// TIA Portal project "EMS" (V15.1) (continued)
   "Carrier_08_G120DStatusWord.3" AT %I762.3 : Bool;   // Bit_03_FAULT
   "Carrier_08_G120DStatusWord.4" AT %I762.4 : Bool;   // Bit_04_OFF2
   "Carrier_08_G120DStatusWord.5" AT %I762.5 : Bool;   // Bit_05_OFF3
   "Carrier_08_G120DStatusWord.6" AT %I762.6 : Bool;   // Bit_06_LOCK_OUT
   "Carrier_08_G120DStatusWord.7" AT %I762.7 : Bool;   // Bit_07_WARN
   "Carrier_08_G120DStatusWord.8" AT %I763.0 : Bool;   // Bit_08_NO_DEVIATION
   "Carrier_08_G120DStatusWord.9" AT %I763.1 : Bool;   // Bit_09_CONTR_PLC
   "Carrier_08_G120DStatusWord.10" AT %I763.2 : Bool;   // Bit_10_F_MAX
   "Carrier_08_G120DStatusWord.11" AT %I763.3 : Bool;   // Bit_11_LIMIT_REACHED
   "Carrier_08_G120DStatusWord.12" AT %I763.4 : Bool;   // Bit_12_BRAKE_OPEN
   "Carrier_08_G120DStatusWord.13" AT %I763.5 : Bool;   // Bit_13_NO_OVERTEMP
   "Carrier_08_G120DStatusWord.14" AT %I763.6 : Bool;   // Bit_14_CW_CCW
   "Carrier_08_G120DStatusWord.15" AT %I763.7 : Bool;   // Bit_15_OVERL
   "Carrier_08_Slot2_Input" AT %IW764 : Word;   // SLOT 2 INPUT WORD
   "Carrier_08_CrashDetectSW" AT %I764.0 : Bool;   // CRASH DETECT SW
   "Carrier_08_SpareSafetyInput(2_1)" AT %I764.1 : Bool;   // SPARE SAFETY INPUT
   "Carrier_08_SpareSafetyInput(2_2)" AT %I764.2 : Bool;   // SPARE SAFETY INPUT
   "Carrier_08_SpareSafetyInput(2_3)" AT %I764.3 : Bool;   // SPARE SAFETY INPUT
   "Carrier_08_SpareSafetyInput(2_4)" AT %I764.4 : Bool;   // SPARE SAFETY INPUT
   "Carrier_08_SpareSafetyInput(2_5)" AT %I764.5 : Bool;   // SPARE SAFETY INPUT
   "Carrier_08_SpareSafetyInput(2_6)" AT %I764.6 : Bool;   // SPARE SAFETY INPUT
   "Carrier_08_SpareSafetyInput(2_7)" AT %I764.7 : Bool;   // SPARE SAFETY INPUT
   "Carrier_08_Slot3_SafetyOutput" AT %IW765 : Word;   // SLOT 3 SAFETY OUTPUT WORD
   "Carrier_08_Crash_Detect_OK" AT %I765.0 : Bool;   // CARRIER CRASH DETECT
   "Carrier_08_SpareSafetyOutput(3_1)" AT %I765.1 : Bool;   // SPARE SAFETY OUTPUT
   "Carrier_08_SpareSafetyOutput(3_2)" AT %I765.2 : Bool;   // SPARE SAFETY OUTPUT
   "Carrier_08_SpareSafetyOutput(3_3)" AT %I765.3 : Bool;   // SPARE SAFETY OUTPUT
   "Carrier_08_SpareSafetyOutput(3_4)" AT %I765.4 : Bool;   // SPARE SAFETY OUTPUT
   "Carrier_08_SpareSafetyOutput(3_5)" AT %I765.5 : Bool;   // SPARE SAFETY OUTPUT
   "Carrier_08_SpareSafetyOutput(3_6)" AT %I765.6 : Bool;   // SPARE SAFETY OUTPUT
   "Carrier_08_SpareSafetyOutput(3_7)" AT %I765.7 : Bool;   // SPARE SAFETY OUTPUT
   "Carrier_08_Slot4_Input" AT %IW766 : Word;   // SLOT 4 INPUT WORD
   "Carrier_08_480VPowerOn_MDCB1" AT %I766.0 : Bool;   // 480 VAC POWER ON MDCB 1
   "Carrier_08_SpareInput(4_1)" AT %I766.1 : Bool;   // SPARE INPUT
   "Carrier_08_SpareInput(4_2)" AT %I766.2 : Bool;   // SPARE INPUT
   "Carrier_08_SitopSelectStatus" AT %I766.3 : Bool;   // SITOP SELECT STATUS
   "Carrier_08_DCsupplyOnPSCB2" AT %I766.4 : Bool;   // DC SUPPLY ON PSCB 2
   "Carrier_08_SpareInput(4_5)" AT %I766.5 : Bool;   // SPARE INPUT
   "Carrier_08_SpareInput(4_6)" AT %I766.6 : Bool;   // SPARE INPUT
   "Carrier_08_SpareInput(4_7)" AT %I766.7 : Bool;   // SPARE INPUT
   "Carrier_08_PB1_ProdHoldLH" AT %I767.0 : Bool;   // PB 1 PRODUCTION HOLD LH
   "Carrier_08_PB2_ResetLH" AT %I767.1 : Bool;   // PB 2 RESET LH
   "Carrier_08_PB3_ProdHoldRH" AT %I767.2 : Bool;   // PB 3 PRODUCTION HOLD RH
   "Carrier_08_PB4_ResetRH" AT %I767.3 : Bool;   // PB 4 RESET RH
   "Carrier_08_SpareInput(4_14)" AT %I767.4 : Bool;   // SPARE INPUT
   "Carrier_08_SpareInput(4_15)" AT %I767.5 : Bool;   // SPARE INPUT
   "Carrier_08_SpareInput(4_16)" AT %I767.6 : Bool;   // SPARE INPUT
   "Carrier_08_SpareInput(4_17)" AT %I767.7 : Bool;   // SPARE INPUT
   "Carrier_08_Slot5_Output" AT %IW768 : Word;   // SLOT 5 OUTPUT WORD
   "Carrier_08_IRD400_HMI_24VDC_ENABLE" AT %I768.0 : Bool;   // IRD 400 PANEL HMI 24V DC POWER
   "Carrier_08_FaultLight_LH" AT %I768.1 : Bool;   // FAULT LIGHT LH
   "Carrier_08_RunLight_LH" AT %I768.2 : Bool;   // RUN LIGHT LH
   "Carrier_08_FaultLight_RH" AT %I768.3 : Bool;   // FAULT LIGHT RH
   "Carrier_08_RunLight_RH" AT %I768.4 : Bool;   // RUN LIGHT RH
   "Carrier_08_SpareOutput(5_5)" AT %I768.5 : Bool;   // SPARE OUTPUT
   "Carrier_08_SpareOutput(5_6)" AT %I768.6 : Bool;   // SPARE OUTPUT
   "Carrier_08_SpareOutput(5_7)" AT %I768.7 : Bool;   // SPARE OUTPUT
   "Carrier_08_ActualSpeed" AT %IW770 : Word;   // ACTUAL SPEED
   "Carrier_08_CarrierDriveAlarm" AT %IW772 : Word;   // CARRIER DRIVE ALARM
   "Carrier_08_CarrierDriveWarning" AT %IW774 : Word;   // CARRIER DRIVE WARNING
   "Carrier_09_Status" AT %IW800 : Word;   // CARRIER STATUS WORD
   "Carrier_09_Status.0" AT %I800.0 : Bool;   // HEARTBEAT
   "Carrier_09_Status.1" AT %I800.1 : Bool;   // MANUAL
   "Carrier_09_Status.2" AT %I800.2 : Bool;   // IN_AUTO
   "Carrier_09_Status.3" AT %I800.3 : Bool;   // POSITIONING_COMPLETE
   "Carrier_09_Status.4" AT %I800.4 : Bool;   // PRODUCTION HOLD
   "Carrier_09_Status.5" AT %I800.5 : Bool;   // CARRIER MOVING FORWARD
   "Carrier_09_Status.6" AT %I800.6 : Bool;   // CARRIER MOVING REVERSE
   "Carrier_09_Status.7" AT %I800.7 : Bool;   // CARRIER FAULT
   "Carrier_09_Status.8" AT %I801.0 : Bool;   // CRASH DETECT TRIPPED
   "Carrier_09_Status.9" AT %I801.1 : Bool;
   "Carrier_09_Status.10" AT %I801.2 : Bool;
   "Carrier_09_Status.11" AT %I801.3 : Bool;
   "Carrier_09_Status.12" AT %I801.4 : Bool;
   "Carrier_09_Status.13" AT %I801.5 : Bool;
   "Carrier_09_Status.14" AT %I801.6 : Bool;
   "Carrier_09_Status.15" AT %I801.7 : Bool;
   "Carrier_09_SDCFaultCode" AT %IW802 : Word;   // SDC FAULT CODE
   "Carrier_09_CarrierPosition" AT %ID804 : DWord;   // CARRIER POSITION
   "Carrier_09_CarrierNumber" AT %IW808 : Word;   // CARRIER NUMBER
   "Carrier_09_G120DControlWord" AT %IW810 : Word;   // G120D_STW1_CONTROL
   "Carrier_09_G120DControlWord.0" AT %I810.0 : Bool;   // Bit_00_ON
   "Carrier_09_G120DControlWord.1" AT %I810.1 : Bool;   // Bit_01_AUS2_INH
   "Carrier_09_G120DControlWord.2" AT %I810.2 : Bool;   // Bit_02_AUS3_STOP
   "Carrier_09_G120DControlWord.3" AT %I810.3 : Bool;   // Bit_03_EN
   "Carrier_09_G120DControlWord.4" AT %I810.4 : Bool;   // Bit_04_EN_RAMP
   "Carrier_09_G120DControlWord.5" AT %I810.5 : Bool;   // Bit_05_START_RAMP
   "Carrier_09_G120DControlWord.6" AT %I810.6 : Bool;   // Bit_06_SETPOINT
   "Carrier_09_G120DControlWord.7" AT %I810.7 : Bool;   // Bit_07_RESET
   "Carrier_09_G120DControlWord.8" AT %I811.0 : Bool;   // Bit_08_JOG_R
   "Carrier_09_G120DControlWord.9" AT %I811.1 : Bool;   // Bit_09_JOG_L
   "Carrier_09_G120DControlWord.10" AT %I811.2 : Bool;   // Bit_10_CONTR_PLC
   "Carrier_09_G120DControlWord.11" AT %I811.3 : Bool;   // Bit_11_REVERSE
   "Carrier_09_G120DControlWord.12" AT %I811.4 : Bool;   // Bit_12_BRAKE_RELEASE
   "Carrier_09_G120DControlWord.13" AT %I811.5 : Bool;   // Bit_13_DDS
   "Carrier_09_G120DControlWord.14" AT %I811.6 : Bool;   // Bit_14_DO0
   "Carrier_09_G120DControlWord.15" AT %I811.7 : Bool;   // Bit_15_DO1
   "Carrier_09_G120DStatusWord" AT %IW812 : Word;   // G120D_ZSW1_STATUS
   "Carrier_09_G120DStatusWord.0" AT %I812.0 : Bool;   // Bit_00_READY_RUN
   "Carrier_09_G120DStatusWord.1" AT %I812.1 : Bool;   // Bit_01_READY_ON
   "Carrier_09_G120DStatusWord.2" AT %I812.2 : Bool;   // Bit_02_ENABLE
   "Carrier_09_G120DStatusWord.3" AT %I812.3 : Bool;   // Bit_03_FAULT
   "Carrier_09_G120DStatusWord.4" AT %I812.4 : Bool;   // Bit_04_OFF2
   "Carrier_09_G120DStatusWord.5" AT %I812.5 : Bool;   // Bit_05_OFF3
   "Carrier_09_G120DStatusWord.6" AT %I812.6 : Bool;   // Bit_06_LOCK_OUT
   "Carrier_09_G120DStatusWord.7" AT %I812.7 : Bool;   // Bit_07_WARN
   "Carrier_09_G120DStatusWord.8" AT %I813.0 : Bool;   // Bit_08_NO_DEVIATION
   "Carrier_09_G120DStatusWord.9" AT %I813.1 : Bool;   // Bit_09_CONTR_PLC
   "Carrier_09_G120DStatusWord.10" AT %I813.2 : Bool;   // Bit_10_F_MAX
   "Carrier_09_G120DStatusWord.11" AT %I813.3 : Bool;   // Bit_11_LIMIT_REACHED
   "Carrier_09_G120DStatusWord.12" AT %I813.4 : Bool;   // Bit_12_BRAKE_OPEN
   "Carrier_09_G120DStatusWord.13" AT %I813.5 : Bool;   // Bit_13_NO_OVERTEMP
   "Carrier_09_G120DStatusWord.14" AT %I813.6 : Bool;   // Bit_14_CW_CCW
   "Carrier_09_G120DStatusWord.15" AT %I813.7 : Bool;   // Bit_15_OVERL
   "Carrier_09_Slot2_Input" AT %IW814 : Word;   // SLOT 2 INPUT WORD
   "Carrier_09_CrashDetectSW" AT %I814.0 : Bool;   // CRASH DETECT SW
   "Carrier_09_SpareSafetyInput(2_1)" AT %I814.1 : Bool;   // SPARE SAFETY INPUT
   "Carrier_09_SpareSafetyInput(2_2)" AT %I814.2 : Bool;   // SPARE SAFETY INPUT
   "Carrier_09_SpareSafetyInput(2_3)" AT %I814.3 : Bool;   // SPARE SAFETY INPUT
   "Carrier_09_SpareSafetyInput(2_4)" AT %I814.4 : Bool;   // SPARE SAFETY INPUT
   "Carrier_09_SpareSafetyInput(2_5)" AT %I814.5 : Bool;   // SPARE SAFETY INPUT
   "Carrier_09_SpareSafetyInput(2_6)" AT %I814.6 : Bool;   // SPARE SAFETY INPUT
   "Carrier_09_SpareSafetyInput(2_7)" AT %I814.7 : Bool;   // SPARE SAFETY INPUT
   "Carrier_09_Slot3_SafetyOutput" AT %IW815 : Word;   // SLOT 3 SAFETY OUTPUT WORD
   "Carrier_09_Crash_Detect_OK" AT %I815.0 : Bool;   // CARRIER CRASH DETECT
   "Carrier_09_SpareSafetyOutput(3_1)" AT %I815.1 : Bool;   // SPARE SAFETY OUTPUT
   "Carrier_09_SpareSafetyOutput(3_2)" AT %I815.2 : Bool;   // SPARE SAFETY OUTPUT
   "Carrier_09_SpareSafetyOutput(3_3)" AT %I815.3 : Bool;   // SPARE SAFETY OUTPUT
   "Carrier_09_SpareSafetyOutput(3_4)" AT %I815.4 : Bool;   // SPARE SAFETY OUTPUT
   "Carrier_09_SpareSafetyOutput(3_5)" AT %I815.5 : Bool;   // SPARE SAFETY OUTPUT
   "Carrier_09_SpareSafetyOutput(3_6)" AT %I815.6 : Bool;   // SPARE SAFETY OUTPUT
   "Carrier_09_SpareSafetyOutput(3_7)" AT %I815.7 : Bool;   // SPARE SAFETY OUTPUT
   "Carrier_09_Slot4_Input" AT %IW816 : Word;   // SLOT 4 INPUT WORD
   "Carrier_09_480VPowerOn_MDCB1" AT %I816.0 : Bool;   // 480 VAC POWER ON MDCB 1
   "Carrier_09_SpareInput(4_1)" AT %I816.1 : Bool;   // SPARE INPUT
   "Carrier_09_SpareInput(4_2)" AT %I816.2 : Bool;   // SPARE INPUT
   "Carrier_09_SitopSelectStatus" AT %I816.3 : Bool;   // SITOP SELECT STATUS
   "Carrier_09_DCsupplyOnPSCB2" AT %I816.4 : Bool;   // DC SUPPLY ON PSCB 2
   "Carrier_09_SpareInput(4_5)" AT %I816.5 : Bool;   // SPARE INPUT
   "Carrier_09_SpareInput(4_6)" AT %I816.6 : Bool;   // SPARE INPUT
   "Carrier_09_SpareInput(4_7)" AT %I816.7 : Bool;   // SPARE INPUT
   "Carrier_09_PB1_ProdHoldLH" AT %I817.0 : Bool;   // PB 1 PRODUCTION HOLD LH
   "Carrier_09_PB2_ResetLH" AT %I817.1 : Bool;   // PB 2 RESET LH
   "Carrier_09_PB3_ProdHoldRH" AT %I817.2 : Bool;   // PB 3 PRODUCTION HOLD RH
   "Carrier_09_PB4_ResetRH" AT %I817.3 : Bool;   // PB 4 RESET RH
   "Carrier_09_SpareInput(4_14)" AT %I817.4 : Bool;   // SPARE INPUT
   "Carrier_09_SpareInput(4_15)" AT %I817.5 : Bool;   // SPARE INPUT
   "Carrier_09_SpareInput(4_16)" AT %I817.6 : Bool;   // SPARE INPUT
   "Carrier_09_SpareInput(4_17)" AT %I817.7 : Bool;   // SPARE INPUT
   "Carrier_09_Slot5_Output" AT %IW818 : Word;   // SLOT 5 OUTPUT WORD
   "Carrier_09_IRD400_HMI_24VDC_ENABLE" AT %I818.0 : Bool;   // IRD 400 PANEL HMI 24V DC POWER
   "Carrier_09_FaultLight_LH" AT %I818.1 : Bool;   // FAULT LIGHT LH
   "Carrier_09_RunLight_LH" AT %I818.2 : Bool;   // RUN LIGHT LH
   "Carrier_09_FaultLight_RH" AT %I818.3 : Bool;   // FAULT LIGHT RH
   "Carrier_09_RunLight_RH" AT %I818.4 : Bool;   // RUN LIGHT RH
   "Carrier_09_SpareOutput(5_5)" AT %I818.5 : Bool;   // SPARE OUTPUT
   "Carrier_09_SpareOutput(5_6)" AT %I818.6 : Bool;   // SPARE OUTPUT
   "Carrier_09_SpareOutput(5_7)" AT %I818.7 : Bool;   // SPARE OUTPUT
   "Carrier_09_ActualSpeed" AT %IW820 : Word;   // ACTUAL SPEED
   "Carrier_09_CarrierDriveAlarm" AT %IW822 : Word;   // CARRIER DRIVE ALARM
   "Carrier_09_CarrierDriveWarning" AT %IW824 : Word;   // CARRIER DRIVE WARNING
   "Carrier_10_Status" AT %IW850 : Word;   // CARRIER STATUS WORD
   "Carrier_10_Status.0" AT %I850.0 : Bool;   // HEARTBEAT
   "Carrier_10_Status.1" AT %I850.1 : Bool;   // MANUAL
   "Carrier_10_Status.2" AT %I850.2 : Bool;   // IN_AUTO
   "Carrier_10_Status.3" AT %I850.3 : Bool;   // POSITIONING_COMPLETE
   "Carrier_10_Status.4" AT %I850.4 : Bool;   // PRODUCTION HOLD
   "Carrier_10_Status.5" AT %I850.5 : Bool;   // CARRIER MOVING FORWARD
   "Carrier_10_Status.6" AT %I850.6 : Bool;   // CARRIER MOVING REVERSE
   "Carrier_10_Status.7" AT %I850.7 : Bool;   // CARRIER FAULT
   "Carrier_10_Status.8" AT %I851.0 : Bool;   // CRASH DETECT TRIPPED
   "Carrier_10_Status.9" AT %I851.1 : Bool;
   "Carrier_10_Status.10" AT %I851.2 : Bool;
   "Carrier_10_Status.11" AT %I851.3 : Bool;
   "Carrier_10_Status.12" AT %I851.4 : Bool;
   "Carrier_10_Status.13" AT %I851.5 : Bool;
   "Carrier_10_Status.14" AT %I851.6 : Bool;
   "Carrier_10_Status.15" AT %I851.7 : Bool;
   "Carrier_10_SDCFaultCode" AT %IW852 : Word;   // SDC FAULT CODE
   "Carrier_10_CarrierPosition" AT %ID854 : DWord;   // CARRIER POSITION
   "Carrier_10_CarrierNumber" AT %IW858 : Word;   // CARRIER NUMBER
   "Carrier_10_G120DControlWord" AT %IW860 : Word;   // G120D_STW1_CONTROL
   "Carrier_10_G120DControlWord.0" AT %I860.0 : Bool;   // Bit_00_ON
   "Carrier_10_G120DControlWord.1" AT %I860.1 : Bool;   // Bit_01_AUS2_INH
   "Carrier_10_G120DControlWord.2" AT %I860.2 : Bool;   // Bit_02_AUS3_STOP
   "Carrier_10_G120DControlWord.3" AT %I860.3 : Bool;   // Bit_03_EN
   "Carrier_10_G120DControlWord.4" AT %I860.4 : Bool;   // Bit_04_EN_RAMP
   "Carrier_10_G120DControlWord.5" AT %I860.5 : Bool;   // Bit_05_START_RAMP
   "Carrier_10_G120DControlWord.6" AT %I860.6 : Bool;   // Bit_06_SETPOINT
   "Carrier_10_G120DControlWord.7" AT %I860.7 : Bool;   // Bit_07_RESET
   "Carrier_10_G120DControlWord.8" AT %I861.0 : Bool;   // Bit_08_JOG_R
   "Carrier_10_G120DControlWord.9" AT %I861.1 : Bool;   // Bit_09_JOG_L
   "Carrier_10_G120DControlWord.10" AT %I861.2 : Bool;   // Bit_10_CONTR_PLC
   "Carrier_10_G120DControlWord.11" AT %I861.3 : Bool;   // Bit_11_REVERSE
   "Carrier_10_G120DControlWord.12" AT %I861.4 : Bool;   // Bit_12_BRAKE_RELEASE
   "Carrier_10_G120DControlWord.13" AT %I861.5 : Bool;   // Bit_13_DDS
   "Carrier_10_G120DControlWord.14" AT %I861.6 : Bool;   // Bit_14_DO0
   "Carrier_10_G120DControlWord.15" AT %I861.7 : Bool;   // Bit_15_DO1
   "Carrier_10_G120DStatusWord" AT %IW862 : Word;   // G120D_ZSW1_STATUS
   "Carrier_10_G120DStatusWord.0" AT %I862.0 : Bool;   // Bit_00_READY_RUN
   "Carrier_10_G120DStatusWord.1" AT %I862.1 : Bool;   // Bit_01_READY_ON
   "Carrier_10_G120DStatusWord.2" AT %I862.2 : Bool;   // Bit_02_ENABLE
   "Carrier_10_G120DStatusWord.3" AT %I862.3 : Bool;   // Bit_03_FAULT
   "Carrier_10_G120DStatusWord.4" AT %I862.4 : Bool;   // Bit_04_OFF2
   "Carrier_10_G120DStatusWord.5" AT %I862.5 : Bool;   // Bit_05_OFF3
   "Carrier_10_G120DStatusWord.6" AT %I862.6 : Bool;   // Bit_06_LOCK_OUT
   "Carrier_10_G120DStatusWord.7" AT %I862.7 : Bool;   // Bit_07_WARN
   "Carrier_10_G120DStatusWord.8" AT %I863.0 : Bool;   // Bit_08_NO_DEVIATION
   "Carrier_10_G120DStatusWord.9" AT %I863.1 : Bool;   // Bit_09_CONTR_PLC
   "Carrier_10_G120DStatusWord.10" AT %I863.2 : Bool;   // Bit_10_F_MAX
   "Carrier_10_G120DStatusWord.11" AT %I863.3 : Bool;   // Bit_11_LIMIT_REACHED
   "Carrier_10_G120DStatusWord.12" AT %I863.4 : Bool;   // Bit_12_BRAKE_OPEN
   "Carrier_10_G120DStatusWord.13" AT %I863.5 : Bool;   // Bit_13_NO_OVERTEMP
   "Carrier_10_G120DStatusWord.14" AT %I863.6 : Bool;   // Bit_14_CW_CCW
   "Carrier_10_G120DStatusWord.15" AT %I863.7 : Bool;   // Bit_15_OVERL
   "Carrier_10_Slot2_Input" AT %IW864 : Word;   // SLOT 2 INPUT WORD
   "Carrier_10_CrashDetectSW" AT %I864.0 : Bool;   // CRASH DETECT SW
   "Carrier_10_SpareSafetyInput(2_1)" AT %I864.1 : Bool;   // SPARE SAFETY INPUT
   "Carrier_10_SpareSafetyInput(2_2)" AT %I864.2 : Bool;   // SPARE SAFETY INPUT
   "Carrier_10_SpareSafetyInput(2_3)" AT %I864.3 : Bool;   // SPARE SAFETY INPUT
   "Carrier_10_SpareSafetyInput(2_4)" AT %I864.4 : Bool;   // SPARE SAFETY INPUT
   "Carrier_10_SpareSafetyInput(2_5)" AT %I864.5 : Bool;   // SPARE SAFETY INPUT
   "Carrier_10_SpareSafetyInput(2_6)" AT %I864.6 : Bool;   // SPARE SAFETY INPUT
   "Carrier_10_SpareSafetyInput(2_7)" AT %I864.7 : Bool;   // SPARE SAFETY INPUT
   "Carrier_10_Slot3_SafetyOutput" AT %IW865 : Word;   // SLOT 3 SAFETY OUTPUT WORD
   "Carrier_10_Crash_Detect_OK" AT %I865.0 : Bool;   // CARRIER CRASH DETECT
   "Carrier_10_SpareSafetyOutput(3_1)" AT %I865.1 : Bool;   // SPARE SAFETY OUTPUT
   "Carrier_10_SpareSafetyOutput(3_2)" AT %I865.2 : Bool;   // SPARE SAFETY OUTPUT
   "Carrier_10_SpareSafetyOutput(3_3)" AT %I865.3 : Bool;   // SPARE SAFETY OUTPUT
   "Carrier_10_SpareSafetyOutput(3_4)" AT %I865.4 : Bool;   // SPARE SAFETY OUTPUT
   "Carrier_10_SpareSafetyOutput(3_5)" AT %I865.5 : Bool;   // SPARE SAFETY OUTPUT
   "Carrier_10_SpareSafetyOutput(3_6)" AT %I865.6 : Bool;   // SPARE SAFETY OUTPUT
   "Carrier_10_SpareSafetyOutput(3_7)" AT %I865.7 : Bool;   // SPARE SAFETY OUTPUT
   "Carrier_10_Slot4_Input" AT %IW866 : Word;   // SLOT 4 INPUT WORD
   "Carrier_10_480VPowerOn_MDCB1" AT %I866.0 : Bool;   // 480 VAC POWER ON MDCB 1
   "Carrier_10_SpareInput(4_1)" AT %I866.1 : Bool;   // SPARE INPUT
   "Carrier_10_SpareInput(4_2)" AT %I866.2 : Bool;   // SPARE INPUT
   "Carrier_10_SitopSelectStatus" AT %I866.3 : Bool;   // SITOP SELECT STATUS
   "Carrier_10_DCsupplyOnPSCB2" AT %I866.4 : Bool;   // DC SUPPLY ON PSCB 2
   "Carrier_10_SpareInput(4_5)" AT %I866.5 : Bool;   // SPARE INPUT
   "Carrier_10_SpareInput(4_6)" AT %I866.6 : Bool;   // SPARE INPUT
   "Carrier_10_SpareInput(4_7)" AT %I866.7 : Bool;   // SPARE INPUT
   "Carrier_10_PB1_ProdHoldLH" AT %I867.0 : Bool;   // PB 1 PRODUCTION HOLD LH
   "Carrier_10_PB2_ResetLH" AT %I867.1 : Bool;   // PB 2 RESET LH
   "Carrier_10_PB3_ProdHoldRH" AT %I867.2 : Bool;   // PB 3 PRODUCTION HOLD RH
   "Carrier_10_PB4_ResetRH" AT %I867.3 : Bool;   // PB 4 RESET RH
   "Carrier_10_SpareInput(4_14)" AT %I867.4 : Bool;   // SPARE INPUT
   "Carrier_10_SpareInput(4_15)" AT %I867.5 : Bool;   // SPARE INPUT
   "Carrier_10_SpareInput(4_16)" AT %I867.6 : Bool;   // SPARE INPUT
   "Carrier_10_SpareInput(4_17)" AT %I867.7 : Bool;   // SPARE INPUT
   "Carrier_10_Slot5_Output" AT %IW868 : Word;   // SLOT 5 OUTPUT WORD
   "Carrier_10_IRD400_HMI_24VDC_ENABLE" AT %I868.0 : Bool;   // IRD 400 PANEL HMI 24V DC POWER
   "Carrier_10_FaultLight_LH" AT %I868.1 : Bool;   // FAULT LIGHT LH
   "Carrier_10_RunLight_LH" AT %I868.2 : Bool;   // RUN LIGHT LH
   "Carrier_10_FaultLight_RH" AT %I868.3 : Bool;   // FAULT LIGHT RH
   "Carrier_10_RunLight_RH" AT %I868.4 : Bool;   // RUN LIGHT RH
   "Carrier_10_SpareOutput(5_5)" AT %I868.5 : Bool;   // SPARE OUTPUT
   "Carrier_10_SpareOutput(5_6)" AT %I868.6 : Bool;   // SPARE OUTPUT
   "Carrier_10_SpareOutput(5_7)" AT %I868.7 : Bool;   // SPARE OUTPUT
   "Carrier_10_ActualSpeed" AT %IW870 : Word;   // ACTUAL SPEED
   "Carrier_10_CarrierDriveAlarm" AT %IW872 : Word;   // CARRIER DRIVE ALARM
   "Carrier_10_CarrierDriveWarning" AT %IW874 : Word;   // CARRIER DRIVE WARNING
   "Carrier_11_Status" AT %IW900 : Word;   // CARRIER STATUS WORD
   "Carrier_11_Status.0" AT %I900.0 : Bool;   // HEARTBEAT
   "Carrier_11_Status.1" AT %I900.1 : Bool;   // MANUAL
   "Carrier_11_Status.2" AT %I900.2 : Bool;   // IN_AUTO
   "Carrier_11_Status.3" AT %I900.3 : Bool;   // POSITIONING_COMPLETE
   "Carrier_11_Status.4" AT %I900.4 : Bool;   // PRODUCTION HOLD
   "Carrier_11_Status.5" AT %I900.5 : Bool;   // CARRIER MOVING FORWARD
   "Carrier_11_Status.6" AT %I900.6 : Bool;   // CARRIER MOVING REVERSE
   "Carrier_11_Status.7" AT %I900.7 : Bool;   // CARRIER FAULT
   "Carrier_11_Status.8" AT %I901.0 : Bool;   // CRASH DETECT TRIPPED
   "Carrier_11_Status.9" AT %I901.1 : Bool;
   "Carrier_11_Status.10" AT %I901.2 : Bool;
   "Carrier_11_Status.11" AT %I901.3 : Bool;
   "Carrier_11_Status.12" AT %I901.4 : Bool;
   "Carrier_11_Status.13" AT %I901.5 : Bool;
   "Carrier_11_Status.14" AT %I901.6 : Bool;
   "Carrier_11_Status.15" AT %I901.7 : Bool;
   "Carrier_11_SDCFaultCode" AT %IW902 : Word;   // SDC FAULT CODE
   "Carrier_11_CarrierPosition" AT %ID904 : DWord;   // CARRIER POSITION
   "Carrier_11_CarrierNumber" AT %IW908 : Word;   // CARRIER NUMBER
   "Carrier_11_G120DControlWord" AT %IW910 : Word;   // G120D_STW1_CONTROL
   "Carrier_11_G120DControlWord.0" AT %I910.0 : Bool;   // Bit_00_ON
   "Carrier_11_G120DControlWord.1" AT %I910.1 : Bool;   // Bit_01_AUS2_INH
   "Carrier_11_G120DControlWord.2" AT %I910.2 : Bool;   // Bit_02_AUS3_STOP
   "Carrier_11_G120DControlWord.3" AT %I910.3 : Bool;   // Bit_03_EN
   "Carrier_11_G120DControlWord.4" AT %I910.4 : Bool;   // Bit_04_EN_RAMP
   "Carrier_11_G120DControlWord.5" AT %I910.5 : Bool;   // Bit_05_START_RAMP
   "Carrier_11_G120DControlWord.6" AT %I910.6 : Bool;   // Bit_06_SETPOINT
   "Carrier_11_G120DControlWord.7" AT %I910.7 : Bool;   // Bit_07_RESET
   "Carrier_11_G120DControlWord.8" AT %I911.0 : Bool;   // Bit_08_JOG_R
   "Carrier_11_G120DControlWord.9" AT %I911.1 : Bool;   // Bit_09_JOG_L
   "Carrier_11_G120DControlWord.10" AT %I911.2 : Bool;   // Bit_10_CONTR_PLC
   "Carrier_11_G120DControlWord.11" AT %I911.3 : Bool;   // Bit_11_REVERSE
   "Carrier_11_G120DControlWord.12" AT %I911.4 : Bool;   // Bit_12_BRAKE_RELEASE
   "Carrier_11_G120DControlWord.13" AT %I911.5 : Bool;   // Bit_13_DDS
   "Carrier_11_G120DControlWord.14" AT %I911.6 : Bool;   // Bit_14_DO0
   "Carrier_11_G120DControlWord.15" AT %I911.7 : Bool;   // Bit_15_DO1
   "Carrier_11_G120DStatusWord" AT %IW912 : Word;   // G120D_ZSW1_STATUS
   "Carrier_11_G120DStatusWord.0" AT %I912.0 : Bool;   // Bit_00_READY_RUN
   "Carrier_11_G120DStatusWord.1" AT %I912.1 : Bool;   // Bit_01_READY_ON
   "Carrier_11_G120DStatusWord.2" AT %I912.2 : Bool;   // Bit_02_ENABLE
   "Carrier_11_G120DStatusWord.3" AT %I912.3 : Bool;   // Bit_03_FAULT
   "Carrier_11_G120DStatusWord.4" AT %I912.4 : Bool;   // Bit_04_OFF2
   "Carrier_11_G120DStatusWord.5" AT %I912.5 : Bool;   // Bit_05_OFF3
   "Carrier_11_G120DStatusWord.6" AT %I912.6 : Bool;   // Bit_06_LOCK_OUT
   "Carrier_11_G120DStatusWord.7" AT %I912.7 : Bool;   // Bit_07_WARN
   "Carrier_11_G120DStatusWord.8" AT %I913.0 : Bool;   // Bit_08_NO_DEVIATION
   "Carrier_11_G120DStatusWord.9" AT %I913.1 : Bool;   // Bit_09_CONTR_PLC
   "Carrier_11_G120DStatusWord.10" AT %I913.2 : Bool;   // Bit_10_F_MAX
   "Carrier_11_G120DStatusWord.11" AT %I913.3 : Bool;   // Bit_11_LIMIT_REACHED
   "Carrier_11_G120DStatusWord.12" AT %I913.4 : Bool;   // Bit_12_BRAKE_OPEN
   "Carrier_11_G120DStatusWord.13" AT %I913.5 : Bool;   // Bit_13_NO_OVERTEMP
   "Carrier_11_G120DStatusWord.14" AT %I913.6 : Bool;   // Bit_14_CW_CCW
   "Carrier_11_G120DStatusWord.15" AT %I913.7 : Bool;   // Bit_15_OVERL
   "Carrier_11_Slot2_Input" AT %IW914 : Word;   // SLOT 2 INPUT WORD
   "Carrier_11_CrashDetectSW" AT %I914.0 : Bool;   // CRASH DETECT SW
   "Carrier_11_SpareSafetyInput(2_1)" AT %I914.1 : Bool;   // SPARE SAFETY INPUT
   "Carrier_11_SpareSafetyInput(2_2)" AT %I914.2 : Bool;   // SPARE SAFETY INPUT
   "Carrier_11_SpareSafetyInput(2_3)" AT %I914.3 : Bool;   // SPARE SAFETY INPUT
   "Carrier_11_SpareSafetyInput(2_4)" AT %I914.4 : Bool;   // SPARE SAFETY INPUT
   "Carrier_11_SpareSafetyInput(2_5)" AT %I914.5 : Bool;   // SPARE SAFETY INPUT
   "Carrier_11_SpareSafetyInput(2_6)" AT %I914.6 : Bool;   // SPARE SAFETY INPUT
   "Carrier_11_SpareSafetyInput(2_7)" AT %I914.7 : Bool;   // SPARE SAFETY INPUT
   "Carrier_11_Slot3_SafetyOutput" AT %IW915 : Word;   // SLOT 3 SAFETY OUTPUT WORD
   "Carrier_11_Crash_Detect_OK" AT %I915.0 : Bool;   // CARRIER CRASH DETECT
   "Carrier_11_SpareSafetyOutput(3_1)" AT %I915.1 : Bool;   // SPARE SAFETY OUTPUT
   "Carrier_11_SpareSafetyOutput(3_2)" AT %I915.2 : Bool;   // SPARE SAFETY OUTPUT
   "Carrier_11_SpareSafetyOutput(3_3)" AT %I915.3 : Bool;   // SPARE SAFETY OUTPUT
   "Carrier_11_SpareSafetyOutput(3_4)" AT %I915.4 : Bool;   // SPARE SAFETY OUTPUT
   "Carrier_11_SpareSafetyOutput(3_5)" AT %I915.5 : Bool;   // SPARE SAFETY OUTPUT
   "Carrier_11_SpareSafetyOutput(3_6)" AT %I915.6 : Bool;   // SPARE SAFETY OUTPUT
   "Carrier_11_SpareSafetyOutput(3_7)" AT %I915.7 : Bool;   // SPARE SAFETY OUTPUT
   "Carrier_11_Slot4_Input" AT %IW916 : Word;   // SLOT 4 INPUT WORD
   "Carrier_11_480VPowerOn_MDCB1" AT %I916.0 : Bool;   // 480 VAC POWER ON MDCB 1
   "Carrier_11_SpareInput(4_1)" AT %I916.1 : Bool;   // SPARE INPUT
   "Carrier_11_SpareInput(4_2)" AT %I916.2 : Bool;   // SPARE INPUT
   "Carrier_11_SitopSelectStatus" AT %I916.3 : Bool;   // SITOP SELECT STATUS
   "Carrier_11_DCsupplyOnPSCB2" AT %I916.4 : Bool;   // DC SUPPLY ON PSCB 2
   "Carrier_11_SpareInput(4_5)" AT %I916.5 : Bool;   // SPARE INPUT
   "Carrier_11_SpareInput(4_6)" AT %I916.6 : Bool;   // SPARE INPUT
   "Carrier_11_SpareInput(4_7)" AT %I916.7 : Bool;   // SPARE INPUT
   "Carrier_11_PB1_ProdHoldLH" AT %I917.0 : Bool;   // PB 1 PRODUCTION HOLD LH
   "Carrier_11_PB2_ResetLH" AT %I917.1 : Bool;   // PB 2 RESET LH
   "Carrier_11_PB3_ProdHoldRH" AT %I917.2 : Bool;   // PB 3 PRODUCTION HOLD RH
   "Carrier_11_PB4_ResetRH" AT %I917.3 : Bool;   // PB 4 RESET RH
   "Carrier_11_SpareInput(4_14)" AT %I917.4 : Bool;   // SPARE INPUT
   "Carrier_11_SpareInput(4_15)" AT %I917.5 : Bool;   // SPARE INPUT
   "Carrier_11_SpareInput(4_16)" AT %I917.6 : Bool;   // SPARE INPUT
   "Carrier_11_SpareInput(4_17)" AT %I917.7 : Bool;   // SPARE INPUT
   "Carrier_11_Slot5_Output" AT %IW918 : Word;   // SLOT 5 OUTPUT WORD
   "Carrier_11_IRD400_HMI_24VDC_ENABLE" AT %I918.0 : Bool;   // IRD 400 PANEL HMI 24V DC POWER
   "Carrier_11_FaultLight_LH" AT %I918.1 : Bool;   // FAULT LIGHT LH
   "Carrier_11_RunLight_LH" AT %I918.2 : Bool;   // RUN LIGHT LH
   "Carrier_11_FaultLight_RH" AT %I918.3 : Bool;   // FAULT LIGHT RH
   "Carrier_11_RunLight_RH" AT %I918.4 : Bool;   // RUN LIGHT RH
   "Carrier_11_SpareOutput(5_5)" AT %I918.5 : Bool;   // SPARE OUTPUT
   "Carrier_11_SpareOutput(5_6)" AT %I918.6 : Bool;   // SPARE OUTPUT
   "Carrier_11_SpareOutput(5_7)" AT %I918.7 : Bool;   // SPARE OUTPUT
   "Carrier_11_ActualSpeed" AT %IW920 : Word;   // ACTUAL SPEED
   "Carrier_11_CarrierDriveAlarm" AT %IW922 : Word;   // CARRIER DRIVE ALARM
   "Carrier_11_CarrierDriveWarning" AT %IW924 : Word;   // CARRIER DRIVE WARNING
   "Carrier_12_Status" AT %IW950 : Word;   // CARRIER STATUS WORD
   "Carrier_12_Status.0" AT %I950.0 : Bool;   // HEARTBEAT
   "Carrier_12_Status.1" AT %I950.1 : Bool;   // MANUAL
   "Carrier_12_Status.2" AT %I950.2 : Bool;   // IN_AUTO
   "Carrier_12_Status.3" AT %I950.3 : Bool;   // POSITIONING_COMPLETE
   "Carrier_12_Status.4" AT %I950.4 : Bool;   // PRODUCTION HOLD
   "Carrier_12_Status.5" AT %I950.5 : Bool;   // CARRIER MOVING FORWARD
   "Carrier_12_Status.6" AT %I950.6 : Bool;   // CARRIER MOVING REVERSE
   "Carrier_12_Status.7" AT %I950.7 : Bool;   // CARRIER FAULT
   "Carrier_12_Status.8" AT %I951.0 : Bool;   // CRASH DETECT TRIPPED
   "Carrier_12_Status.9" AT %I951.1 : Bool;
   "Carrier_12_Status.10" AT %I951.2 : Bool;
   "Carrier_12_Status.11" AT %I951.3 : Bool;
   "Carrier_12_Status.12" AT %I951.4 : Bool;
   "Carrier_12_Status.13" AT %I951.5 : Bool;
   "Carrier_12_Status.14" AT %I951.6 : Bool;
   "Carrier_12_Status.15" AT %I951.7 : Bool;
   "Carrier_12_SDCFaultCode" AT %IW952 : Word;   // SDC FAULT CODE
   "Carrier_12_CarrierPosition" AT %ID954 : DWord;   // CARRIER POSITION
   "Carrier_12_CarrierNumber" AT %IW958 : Word;   // CARRIER NUMBER
   "Carrier_12_G120DControlWord" AT %IW960 : Word;   // G120D_STW1_CONTROL
   "Carrier_12_G120DControlWord.0" AT %I960.0 : Bool;   // Bit_00_ON
   "Carrier_12_G120DControlWord.1" AT %I960.1 : Bool;   // Bit_01_AUS2_INH
   "Carrier_12_G120DControlWord.2" AT %I960.2 : Bool;   // Bit_02_AUS3_STOP
   "Carrier_12_G120DControlWord.3" AT %I960.3 : Bool;   // Bit_03_EN
   "Carrier_12_G120DControlWord.4" AT %I960.4 : Bool;   // Bit_04_EN_RAMP
   "Carrier_12_G120DControlWord.5" AT %I960.5 : Bool;   // Bit_05_START_RAMP
   "Carrier_12_G120DControlWord.6" AT %I960.6 : Bool;   // Bit_06_SETPOINT
   "Carrier_12_G120DControlWord.7" AT %I960.7 : Bool;   // Bit_07_RESET
   "Carrier_12_G120DControlWord.8" AT %I961.0 : Bool;   // Bit_08_JOG_R
   "Carrier_12_G120DControlWord.9" AT %I961.1 : Bool;   // Bit_09_JOG_L
   "Carrier_12_G120DControlWord.10" AT %I961.2 : Bool;   // Bit_10_CONTR_PLC
   "Carrier_12_G120DControlWord.11" AT %I961.3 : Bool;   // Bit_11_REVERSE
   "Carrier_12_G120DControlWord.12" AT %I961.4 : Bool;   // Bit_12_BRAKE_RELEASE
   "Carrier_12_G120DControlWord.13" AT %I961.5 : Bool;   // Bit_13_DDS
   "Carrier_12_G120DControlWord.14" AT %I961.6 : Bool;   // Bit_14_DO0
   "Carrier_12_G120DControlWord.15" AT %I961.7 : Bool;   // Bit_15_DO1
   "Carrier_12_G120DStatusWord" AT %IW962 : Word;   // G120D_ZSW1_STATUS
   "Carrier_12_G120DStatusWord.0" AT %I962.0 : Bool;   // Bit_00_READY_RUN
   "Carrier_12_G120DStatusWord.1" AT %I962.1 : Bool;   // Bit_01_READY_ON
   "Carrier_12_G120DStatusWord.2" AT %I962.2 : Bool;   // Bit_02_ENABLE
   "Carrier_12_G120DStatusWord.3" AT %I962.3 : Bool;   // Bit_03_FAULT
   "Carrier_12_G120DStatusWord.4" AT %I962.4 : Bool;   // Bit_04_OFF2
   "Carrier_12_G120DStatusWord.5" AT %I962.5 : Bool;   // Bit_05_OFF3
   "Carrier_12_G120DStatusWord.6" AT %I962.6 : Bool;   // Bit_06_LOCK_OUT
   "Carrier_12_G120DStatusWord.7" AT %I962.7 : Bool;   // Bit_07_WARN
   "Carrier_12_G120DStatusWord.8" AT %I963.0 : Bool;   // Bit_08_NO_DEVIATION
   "Carrier_12_G120DStatusWord.9" AT %I963.1 : Bool;   // Bit_09_CONTR_PLC
   "Carrier_12_G120DStatusWord.10" AT %I963.2 : Bool;   // Bit_10_F_MAX
   "Carrier_12_G120DStatusWord.11" AT %I963.3 : Bool;   // Bit_11_LIMIT_REACHED
   "Carrier_12_G120DStatusWord.12" AT %I963.4 : Bool;   // Bit_12_BRAKE_OPEN
   "Carrier_12_G120DStatusWord.13" AT %I963.5 : Bool;   // Bit_13_NO_OVERTEMP
   "Carrier_12_G120DStatusWord.14" AT %I963.6 : Bool;   // Bit_14_CW_CCW
   "Carrier_12_G120DStatusWord.15" AT %I963.7 : Bool;   // Bit_15_OVERL
   "Carrier_12_Slot2_Input" AT %IW964 : Word;   // SLOT 2 INPUT WORD
   "Carrier_12_CrashDetectSW" AT %I964.0 : Bool;   // CRASH DETECT SW
   "Carrier_12_SpareSafetyInput(2_1)" AT %I964.1 : Bool;   // SPARE SAFETY INPUT
   "Carrier_12_SpareSafetyInput(2_2)" AT %I964.2 : Bool;   // SPARE SAFETY INPUT
   "Carrier_12_SpareSafetyInput(2_3)" AT %I964.3 : Bool;   // SPARE SAFETY INPUT
   "Carrier_12_SpareSafetyInput(2_4)" AT %I964.4 : Bool;   // SPARE SAFETY INPUT
   "Carrier_12_SpareSafetyInput(2_5)" AT %I964.5 : Bool;   // SPARE SAFETY INPUT
   "Carrier_12_SpareSafetyInput(2_6)" AT %I964.6 : Bool;   // SPARE SAFETY INPUT
   "Carrier_12_SpareSafetyInput(2_7)" AT %I964.7 : Bool;   // SPARE SAFETY INPUT
   "Carrier_12_Slot3_SafetyOutput" AT %IW965 : Word;   // SLOT 3 SAFETY OUTPUT WORD
   "Carrier_12_Crash_Detect_OK" AT %I965.0 : Bool;   // CARRIER CRASH DETECT
   "Carrier_12_SpareSafetyOutput(3_1)" AT %I965.1 : Bool;   // SPARE SAFETY OUTPUT
   "Carrier_12_SpareSafetyOutput(3_2)" AT %I965.2 : Bool;   // SPARE SAFETY OUTPUT
   "Carrier_12_SpareSafetyOutput(3_3)" AT %I965.3 : Bool;   // SPARE SAFETY OUTPUT
   "Carrier_12_SpareSafetyOutput(3_4)" AT %I965.4 : Bool;   // SPARE SAFETY OUTPUT
   "Carrier_12_SpareSafetyOutput(3_5)" AT %I965.5 : Bool;   // SPARE SAFETY OUTPUT
   "Carrier_12_SpareSafetyOutput(3_6)" AT %I965.6 : Bool;   // SPARE SAFETY OUTPUT
   "Carrier_12_SpareSafetyOutput(3_7)" AT %I965.7 : Bool;   // SPARE SAFETY OUTPUT
   "Carrier_12_Slot4_Input" AT %IW966 : Word;   // SLOT 4 INPUT WORD
   "Carrier_12_480VPowerOn_MDCB1" AT %I966.0 : Bool;   // 480 VAC POWER ON MDCB 1
   "Carrier_12_SpareInput(4_1)" AT %I966.1 : Bool;   // SPARE INPUT
   "Carrier_12_SpareInput(4_2)" AT %I966.2 : Bool;   // SPARE INPUT
   "Carrier_12_SitopSelectStatus" AT %I966.3 : Bool;   // SITOP SELECT STATUS
   "Carrier_12_DCsupplyOnPSCB2" AT %I966.4 : Bool;   // DC SUPPLY ON PSCB 2
   "Carrier_12_SpareInput(4_5)" AT %I966.5 : Bool;   // SPARE INPUT
   "Carrier_12_SpareInput(4_6)" AT %I966.6 : Bool;   // SPARE INPUT
   "Carrier_12_SpareInput(4_7)" AT %I966.7 : Bool;   // SPARE INPUT
   "Carrier_12_PB1_ProdHoldLH" AT %I967.0 : Bool;   // PB 1 PRODUCTION HOLD LH
   "Carrier_12_PB2_ResetLH" AT %I967.1 : Bool;   // PB 2 RESET LH
   "Carrier_12_PB3_ProdHoldRH" AT %I967.2 : Bool;   // PB 3 PRODUCTION HOLD RH
   "Carrier_12_PB4_ResetRH" AT %I967.3 : Bool;   // PB 4 RESET RH
   "Carrier_12_SpareInput(4_14)" AT %I967.4 : Bool;   // SPARE INPUT
   "Carrier_12_SpareInput(4_15)" AT %I967.5 : Bool;   // SPARE INPUT
   "Carrier_12_SpareInput(4_16)" AT %I967.6 : Bool;   // SPARE INPUT
   "Carrier_12_SpareInput(4_17)" AT %I967.7 : Bool;   // SPARE INPUT
   "Carrier_12_Slot5_Output" AT %IW968 : Word;   // SLOT 5 OUTPUT WORD
   "Carrier_12_IRD400_HMI_24VDC_ENABLE" AT %I968.0 : Bool;   // IRD 400 PANEL HMI 24V DC POWER
   "Carrier_12_FaultLight_LH" AT %I968.1 : Bool;   // FAULT LIGHT LH
   "Carrier_12_RunLight_LH" AT %I968.2 : Bool;   // RUN LIGHT LH
   "Carrier_12_FaultLight_RH" AT %I968.3 : Bool;   // FAULT LIGHT RH
   "Carrier_12_RunLight_RH" AT %I968.4 : Bool;   // RUN LIGHT RH
   "Carrier_12_SpareOutput(5_5)" AT %I968.5 : Bool;   // SPARE OUTPUT
   "Carrier_12_SpareOutput(5_6)" AT %I968.6 : Bool;   // SPARE OUTPUT
   "Carrier_12_SpareOutput(5_7)" AT %I968.7 : Bool;   // SPARE OUTPUT
   "Carrier_12_ActualSpeed" AT %IW970 : Word;   // ACTUAL SPEED
   "Carrier_12_CarrierDriveAlarm" AT %IW972 : Word;   // CARRIER DRIVE ALARM
   "Carrier_12_CarrierDriveWarning" AT %IW974 : Word;   // CARRIER DRIVE WARNING
